		IF ShuttleCarInOut.xPosLimitCatch THEN
			ShuttleCarInOut.xCW:=0;
			ShuttleCarInOut.xMDIDone:=0;
		END_IF;

		IF ShuttleCarInOut.xNegLimitCatch THEN
			ShuttleCarInOut.xCCW:=0;
			ShuttleCarInOut.xMDIDone:=0;
		END_IF;
		ELSE
		ShuttleCarInOut.xCW:=0;
		ShuttleCarInOut.xCCW:=0;
		ShuttleCarInOut.xMDIDone:=0;
	  END_IF;
	END_IF;
	ELSE  (*无就绪信号   或急停的情况下*)
		ShuttleCarInOut.xCW:=0;
		ShuttleCarInOut.xCCW:=0;	
END_IF;
    (*抱闸延时*)
m_tonBrakeDelay(IN:= ShuttleCarInOut.xCW OR ShuttleCarInOut.xCCW,
                                    PT:= ShuttleCarInOut.tBrakeDelay,
                                    Q:=ShuttleCarInOut.xBrake ,
                                    ET:= m_tBrakeDelayCurrentTime);

(*自动上电后把当前位置清零，防止穿梭车不在开关位置*)
IF LDP(TRUE,g_xAuto) THEN
	ShuttleCarInOut.iCurrentPos:=0;
END_IF;
IF ShuttleCarInOut.xCW OR ShuttleCarInOut.xCCW THEN
	ShuttleCarInOut.xBusy:=1;
	ELSE
	ShuttleCarInout.xBusy:=0;
END_IF;

(*暂停，带延时减速斜坡，ShuttleCarInOut.xPauseRamp为减速斜坡输出位*)
m_tonPauseDelay(IN:=g_xPause,PT:= T#2s ,Q:=ShuttleCarInOut.xPauseRamp,ET:= m_tPauseDelayCurrentTime );
IF ShuttleCarInOut.xPauseRamp THEN
	ShuttleCarInOut.xCW:=0;
	ShuttleCarInOut.xCCW:=0;
	ShuttleCarInOut.xBrake:=0;
END_IF;
(*超时报警*)
m_tonOvertimeAlarm(IN:= ShuttleCarInOut.xMDIExe AND (ShuttleCarInOut.iCurrentPos<>ShuttleCarInOut.iDestinationPos) ,
                                           PT:= ShuttleCarInOut.tSetOverTime,
                                           Q:= ShuttleCarInOut.xOvertimeAlarm ,
                                           ET:= m_tOvertimeCurrentTime );
END_FUNCTION_BLOCK

FUNCTION_BLOCK BarCylinder
VAR_IN_OUT
  BarCylinderIO : BarCylinderIO;
END_VAR
VAR
  m_xInitial : BOOL;  (* 初始化 *)
  m_tonLoadDelay : TON;  (* 上料延时 *)
  m_xLoadDelay : BOOL;  (* 上料延时标志位 *)
  m_tLoadDelayCurrentTime : TIME;  (* 上料延时当前时间 *)
END_VAR
  (***********************************************************************
阻挡器模块，
由一个行程开关，一个阻挡器，一个倍速链输送电机组成
具有手动与自动模式
xEmpty显示当前为空料的状态
xUnload为卸料信号，连接下一设备的xEmpty信号
增加分料气缸xBarCylinderSecondary
增加复位功能，Unload NextRun  Empty 能形成死锁，如果Unload 信号一直给，会造成无法复位
*************************************************************************)

IF NOT m_xInitial THEN
	BarCylinderIO.tLoadDelay:=T#3s;
	m_xInitial:=1;
END_IF;
IF g_xManual THEN    (*手动*)
	BarCylinderIO.xNextRun:=0;
	BarCylinderIO.xBarCylinder:=BarCylinderIO.xBarCylinderButton;
	BarCylinderIO.xBarCylinderSecondary	:=BarCylinderIO.xBarSecondaryButton;
	BarCylinderIO.xTransportMotorCW:= BarCylinderIO.xTransportMotorCWButton 
																	AND NOT BarCylinderIO.xTransportMotorCCWButton 
																	AND NOT BarCylinderIO.xTransportMotorCCW ;
	BarCylinderIO.xTransportMotorCCW:=BarCylinderIO.xTransportMotorCCWButton 
																		AND NOT BarCylinderIO.xTransportMotorCWButton 
																		AND NOT BarCylinderIO.xTransportMotorCW;
END_IF;
IF g_xAuto THEN(*自动*)
    IF BarCylinderIO.xUnload   (*下料*)
    	AND NOT BarCylinderIO.xEmpty  (*有料*)
    	AND NOT BarCylinderIO.xNextRun  (*下段线体旋转*)
    	AND NOT (g_xResetSingle AND BarCylinderIO.iDeviceID=g_iDeviceIDSelect)(*无复位信号*)
    	THEN(*收到卸料命令，当阻挡器不为空时*)
    	BarCylinderIO.xBarCylinder:=1;
    	BarCylinderIO.xNextRun:=1;(*确保下料命令只执行一次，防止物料在输送过程中又有卸料命令导致多次卸料*)
    	BarCylinderIO.xTransportMotorCW:=1;
    END_IF;
    IF NOT  BarCylinderIO.xUnload  THEN
    	BarCylinderIO.xNextRun:=0;
    	BarCylinderIO.xBarCylinder:=0;
    END_IF;
    m_tonLoadDelay(IN:= BarCylinderIO.xPresentSwitch ,PT:= BarCylinderIO.tLoadDelay ,Q:= m_xLoadDelay,ET:= m_tLoadDelayCurrentTime );
    IF m_xLoadDelay OR  BarCylinderIO.xNextRun  THEN
    	BarCylinderIO.xEmpty:=0;
    	BarCylinderIO.xBarCylinderSecondary:=1;
    ELSE
    	BarCylinderIO.xEmpty:=1;
    	BarCylinderIO.xBarCylinderSecondary:=0;
    END_IF;
    (*如果为空，气缸顶起*)
   IF  BarCylinderIO.xEmpty  THEN
   	   BarCylinderIO.xBarCylinder:=0;
   END_IF;
   	IF BarCylinderIO.xLoad AND BarCylinderIO.xEmpty  THEN
		BarCylinderIO.xTransportMotorCW:=1;
   	END_IF;  
   	IF (BarCylinderIO.xLoad=0 OR BarCylinderIO.xEmpty=0)  AND (BarCylinderIO.xUnload=0 OR BarCylinderIO.xEmpty) THEN
   		BarCylinderIO.xTransportMotorCW:=0;
   	END_IF;
END_IF;  
IF BarCylinderIO.xEmpty AND BarCylinderIO.xLoad=0 THEN
	BarCylinderIO.iProductCategory:=0;
END_IF;

IF NOT g_xEStop THEN
	 BarCylinderIO.xTransportMotorCW:=0;
	 BarCylinderIO.xTransportMotorCCW:=0;
	 BarCylinderIO.xBarCylinder:=0;
END_IF;

(*//复位*)
IF  (g_xResetSingle AND BarCylinderIO.iDeviceID=g_iDeviceIDSelect)THEN   (* //非正常情况下切断xNextRun不会复位，通过这个标志位会出发报警*)(*增加单体复位*)
	 BarCylinderIO.xNextRun:=0; 
END_IF;
END_FUNCTION_BLOCK
